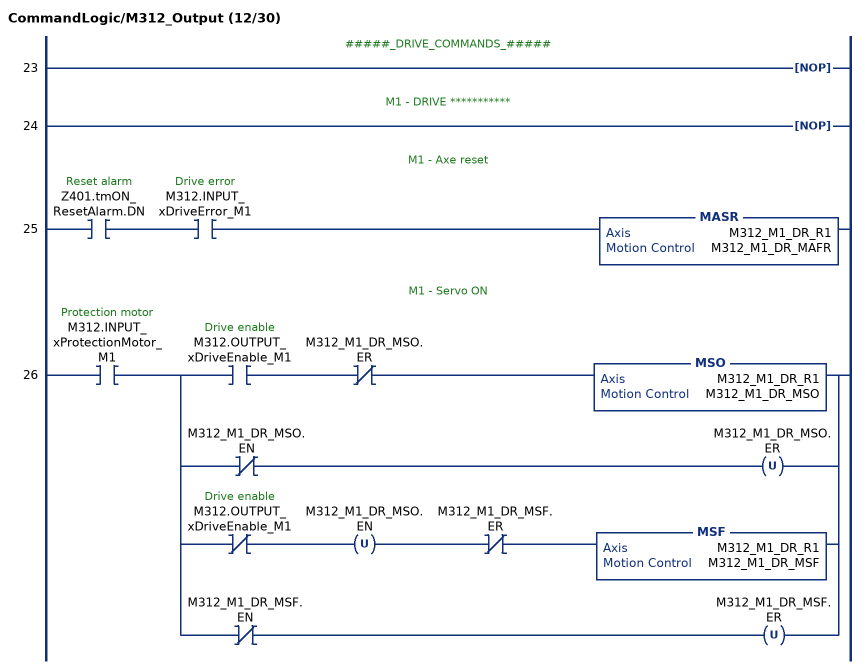
   // #####_DRIVE_COMMANDS_#####
   23: NOP();
   // M1 - DRIVE ***********
   24: NOP();
   // M1 - Axe reset
   25: XIC(Z401.tmON_ResetAlarm.DN)XIC(M312.INPUT_xDriveError_M1)MASR(M312_M1_DR_R1,M312_M1_DR_MAFR);
   // M1 - Servo ON
   26: XIC(M312.INPUT_xProtectionMotor_M1)[XIC(M312.OUTPUT_xDriveEnable_M1) XIO(M312_M1_DR_MSO.ER) MSO(M312_M1_DR_R1,M312_M1_DR_MSO) ,XIO(M312_M1_DR_MSO.EN) OTU(M312_M1_DR_MSO.ER) ,XIO(M312.OUTPUT_xDriveEnable_M1) OTU(M312_M1_DR_MSO.EN) XIO(M312_M1_DR_MSF.ER) MSF(M312_M1_DR_R1,M312_M1_DR_MSF) ,XIO(M312_M1_DR_MSF.EN) OTU(M312_M1_DR_MSF.ER) ];
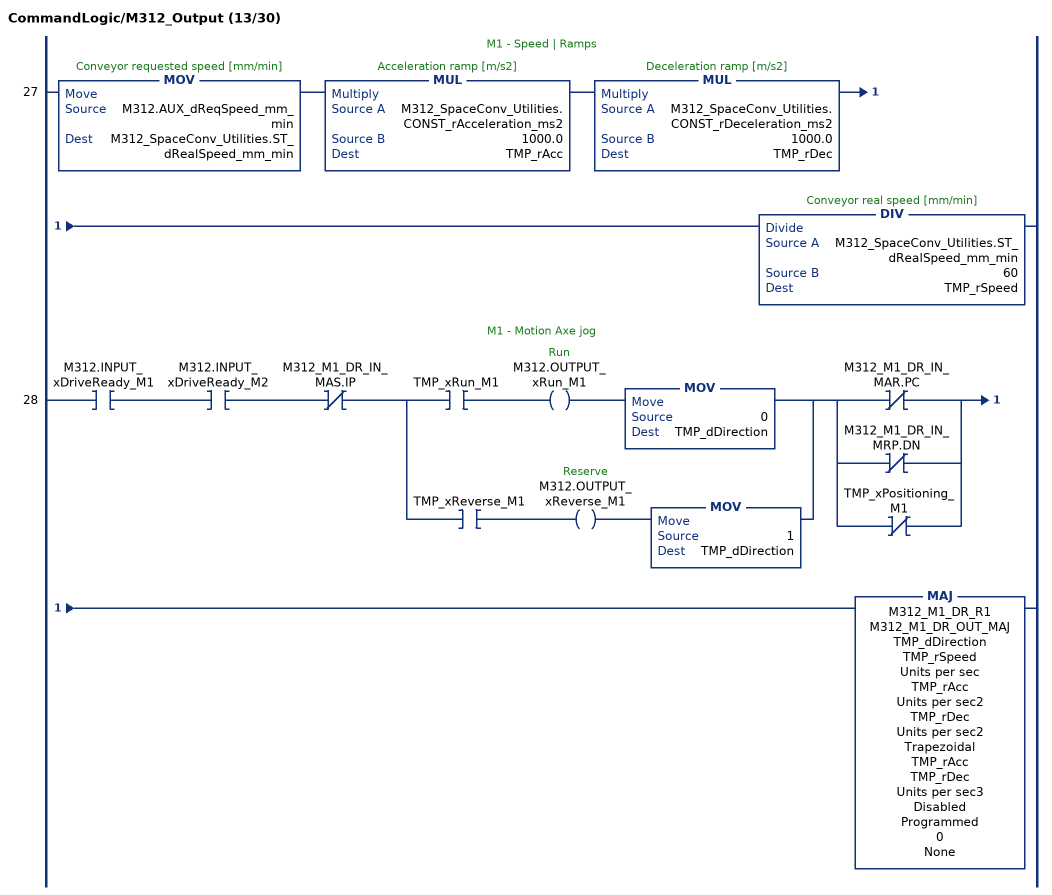
   // M1 - Speed | Ramps
   27: MOV(M312.AUX_dReqSpeed_mm_min,M312_SpaceConv_Utilities.ST_dRealSpeed_mm_min)MUL(M312_SpaceConv_Utilities.CONST_rAcceleration_ms2,1000.0,TMP_rAcc)MUL(M312_SpaceConv_Utilities.CONST_rDeceleration_ms2,1000.0,TMP_rDec)DIV(M312_SpaceConv_Utilities.ST_dRealSpeed_mm_min,60,TMP_rSpeed);
   // M1 - Motion Axe jog
   28: XIC(M312.INPUT_xDriveReady_M1)XIC(M312.INPUT_xDriveReady_M2)XIO(M312_M1_DR_IN_MAS.IP)[XIC(TMP_xRun_M1) OTE(M312.OUTPUT_xRun_M1) MOV(0,TMP_dDirection) ,XIC(TMP_xReverse_M1) OTE(M312.OUTPUT_xReverse_M1) MOV(1,TMP_dDirection) ][XIO(M312_M1_DR_IN_MAR.PC) ,XIO(M312_M1_DR_IN_MRP.DN) ,XIO(TMP_xPositioning_M1) ]MAJ(M312_M1_DR_R1,M312_M1_DR_OUT_MAJ,TMP_dDirection,TMP_rSpeed,Units per sec,TMP_rAcc,Units per sec2,TMP_rDec,Units per sec2,Trapezoidal,TMP_rAcc,TMP_rDec,Units per sec3,Disabled,Programmed,0,None);
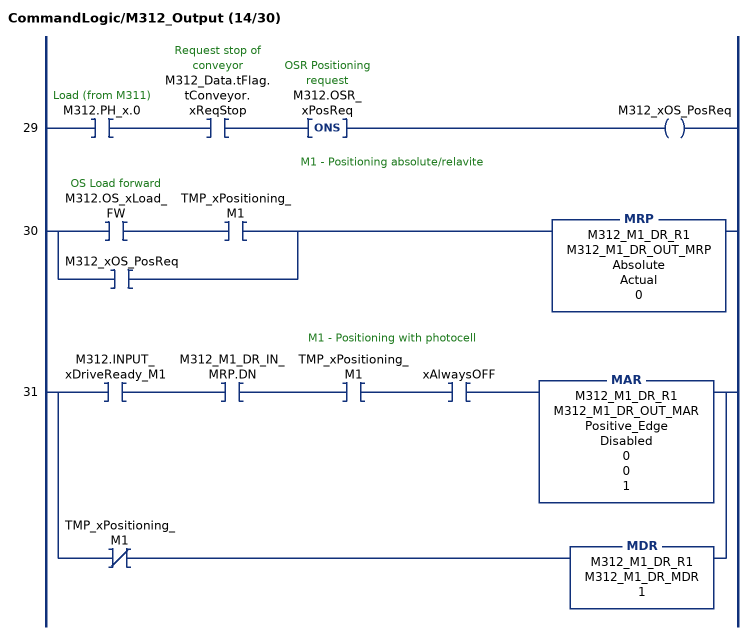
   29: XIC(M312.PH_x.0)XIC(M312_Data.tFlag.tConveyor.xReqStop)ONS(M312.OSR_xPosReq)OTE(M312_xOS_PosReq);
   // M1 - Positioning absolute/relavite
   30: [XIC(M312.OS_xLoad_FW) XIC(TMP_xPositioning_M1) ,XIC(M312_xOS_PosReq) ]MRP(M312_M1_DR_R1,M312_M1_DR_OUT_MRP,Absolute,Actual,0);
   // M1 - Positioning with photocell
   31: [XIC(M312.INPUT_xDriveReady_M1) XIC(M312_M1_DR_IN_MRP.DN) XIC(TMP_xPositioning_M1) XIC(xAlwaysOFF) MAR(M312_M1_DR_R1,M312_M1_DR_OUT_MAR,Positive_Edge,Disabled,0,0,1) ,XIO(TMP_xPositioning_M1) MDR(M312_M1_DR_R1,M312_M1_DR_MDR,1) ];
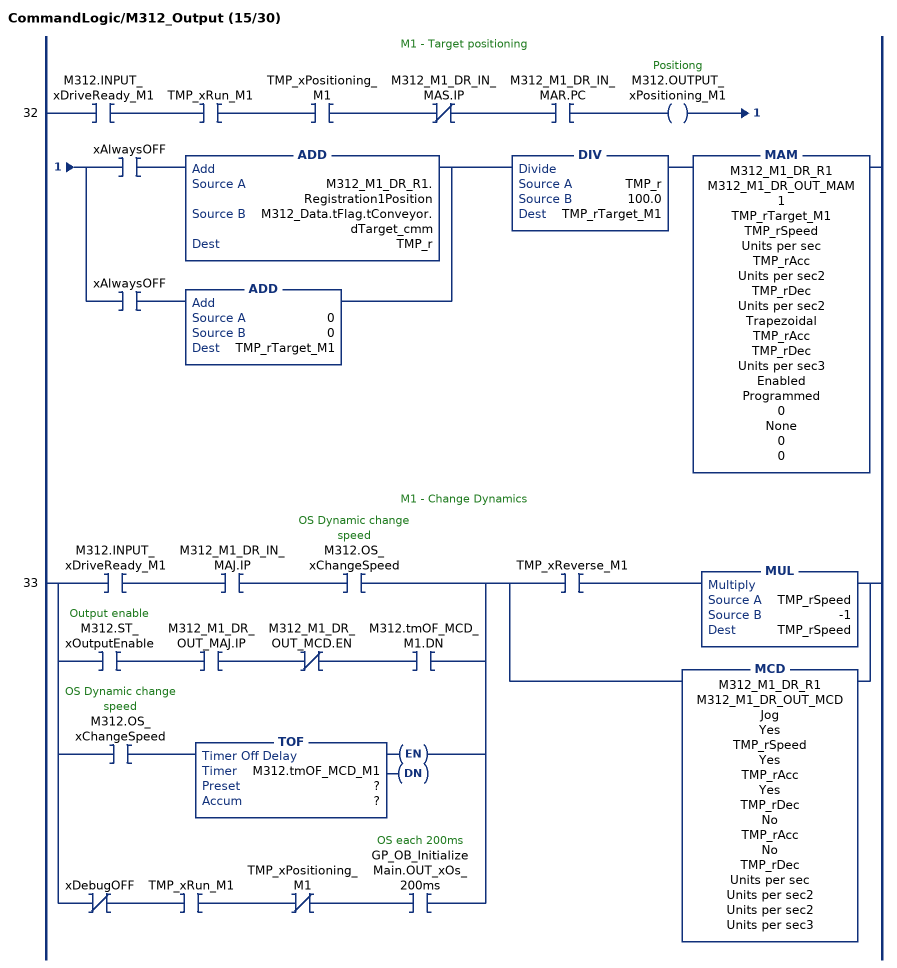
   // M1 - Target positioning
   32: XIC(M312.INPUT_xDriveReady_M1)XIC(TMP_xRun_M1)XIC(TMP_xPositioning_M1)XIO(M312_M1_DR_IN_MAS.IP)XIC(M312_M1_DR_IN_MAR.PC)OTE(M312.OUTPUT_xPositioning_M1)[XIC(xAlwaysOFF) ADD(M312_M1_DR_R1.Registration1Position,M312_Data.tFlag.tConveyor.dTarget_cmm,TMP_r) ,XIC(xAlwaysOFF) ADD(0,0,TMP_rTarget_M1) ]DIV(TMP_r,100.0,TMP_rTarget_M1)MAM(M312_M1_DR_R1,M312_M1_DR_OUT_MAM,1,TMP_rTarget_M1,TMP_rSpeed,Units per sec,TMP_rAcc,Units per sec2,TMP_rDec,Units per sec2,Trapezoidal,TMP_rAcc,TMP_rDec,Units per sec3,Enabled,Programmed,0,None,0,0);
   // M1 - Change Dynamics
   33: [XIC(M312.INPUT_xDriveReady_M1) XIC(M312_M1_DR_IN_MAJ.IP) XIC(M312.OS_xChangeSpeed) ,XIC(M312.ST_xOutputEnable) XIC(M312_M1_DR_OUT_MAJ.IP) XIO(M312_M1_DR_OUT_MCD.EN) XIC(M312.tmOF_MCD_M1.DN) ,XIC(M312.OS_xChangeSpeed) TOF(M312.tmOF_MCD_M1,?,?) ,XIO(xDebugOFF) XIC(TMP_xRun_M1) XIO(TMP_xPositioning_M1) XIC(GP_OB_InitializeMain.OUT_xOs_200ms) ][XIC(TMP_xReverse_M1) MUL(TMP_rSpeed,-1,TMP_rSpeed) ,MCD(M312_M1_DR_R1,M312_M1_DR_OUT_MCD,Jog,Yes,TMP_rSpeed,Yes,TMP_rAcc,Yes,TMP_rDec,No,TMP_rAcc,No,TMP_rDec,Units per sec,Units per sec2,Units per sec2,Units per sec3) ];
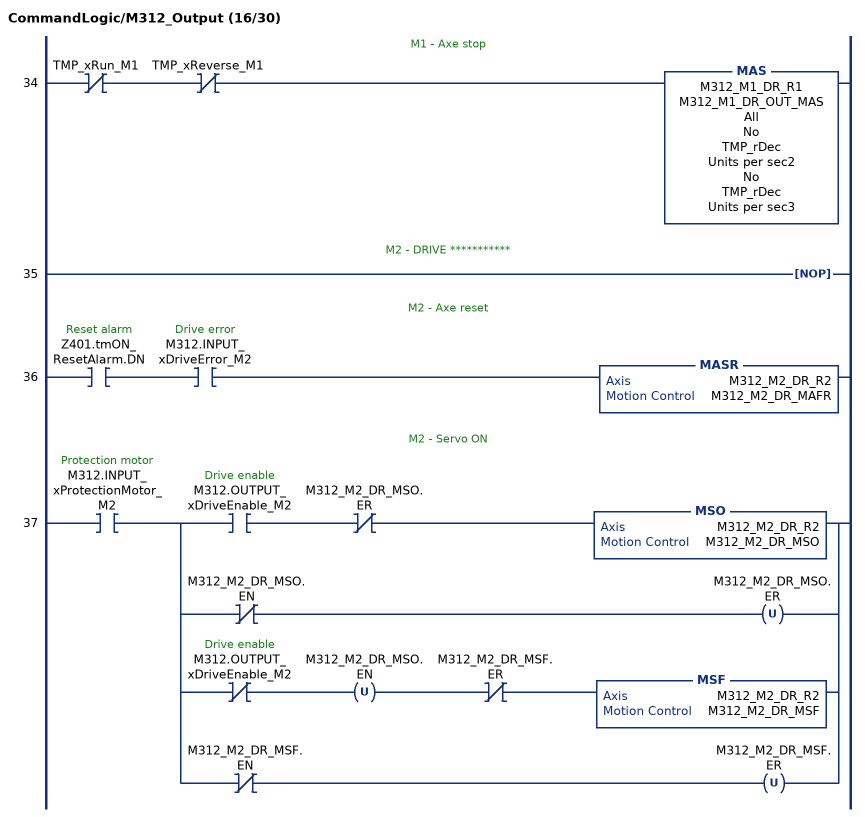
   // M1 - Axe stop
   34: XIO(TMP_xRun_M1)XIO(TMP_xReverse_M1)MAS(M312_M1_DR_R1,M312_M1_DR_OUT_MAS,All,No,TMP_rDec,Units per sec2,No,TMP_rDec,Units per sec3);
   // M2 - DRIVE ***********
   35: NOP();
   // M2 - Axe reset
   36: XIC(Z401.tmON_ResetAlarm.DN)XIC(M312.INPUT_xDriveError_M2)MASR(M312_M2_DR_R2,M312_M2_DR_MAFR);
   // M2 - Servo ON
   37: XIC(M312.INPUT_xProtectionMotor_M2)[XIC(M312.OUTPUT_xDriveEnable_M2) XIO(M312_M2_DR_MSO.ER) MSO(M312_M2_DR_R2,M312_M2_DR_MSO) ,XIO(M312_M2_DR_MSO.EN) OTU(M312_M2_DR_MSO.ER) ,XIO(M312.OUTPUT_xDriveEnable_M2) OTU(M312_M2_DR_MSO.EN) XIO(M312_M2_DR_MSF.ER) MSF(M312_M2_DR_R2,M312_M2_DR_MSF) ,XIO(M312_M2_DR_MSF.EN) OTU(M312_M2_DR_MSF.ER) ];
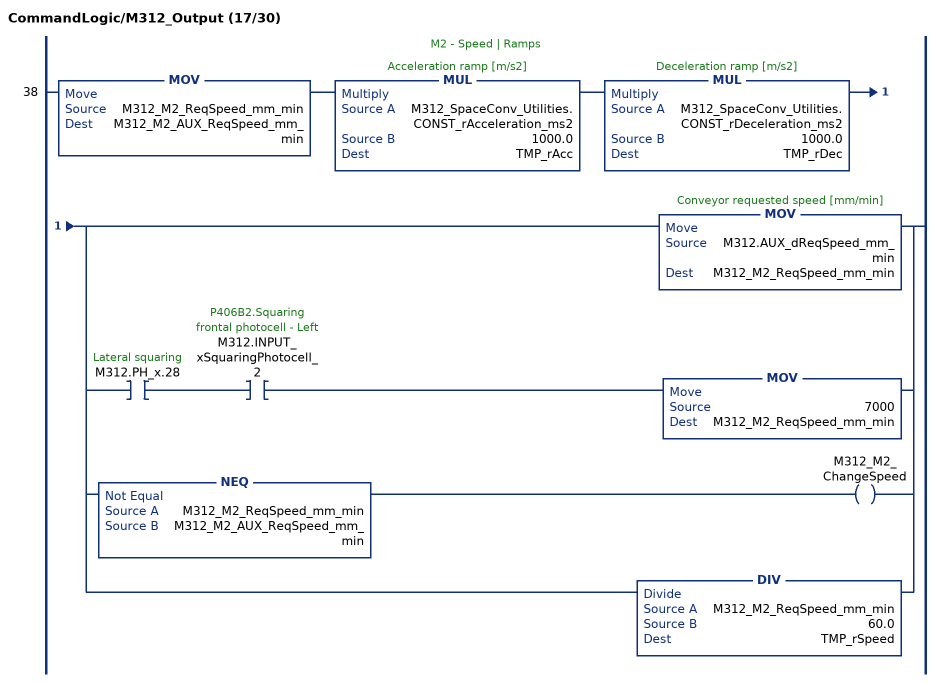
   // M2 - Speed | Ramps
   38: MOV(M312_M2_ReqSpeed_mm_min,M312_M2_AUX_ReqSpeed_mm_min)MUL(M312_SpaceConv_Utilities.CONST_rAcceleration_ms2,1000.0,TMP_rAcc)MUL(M312_SpaceConv_Utilities.CONST_rDeceleration_ms2,1000.0,TMP_rDec)[MOV(M312.AUX_dReqSpeed_mm_min,M312_M2_ReqSpeed_mm_min) ,XIC(M312.PH_x.28) XIC(M312.INPUT_xSquaringPhotocell_2) MOV(7000,M312_M2_ReqSpeed_mm_min) ,NEQ(M312_M2_ReqSpeed_mm_min,M312_M2_AUX_ReqSpeed_mm_min) OTE(M312_M2_ChangeSpeed) ,DIV(M312_M2_ReqSpeed_mm_min,60.0,TMP_rSpeed) ];
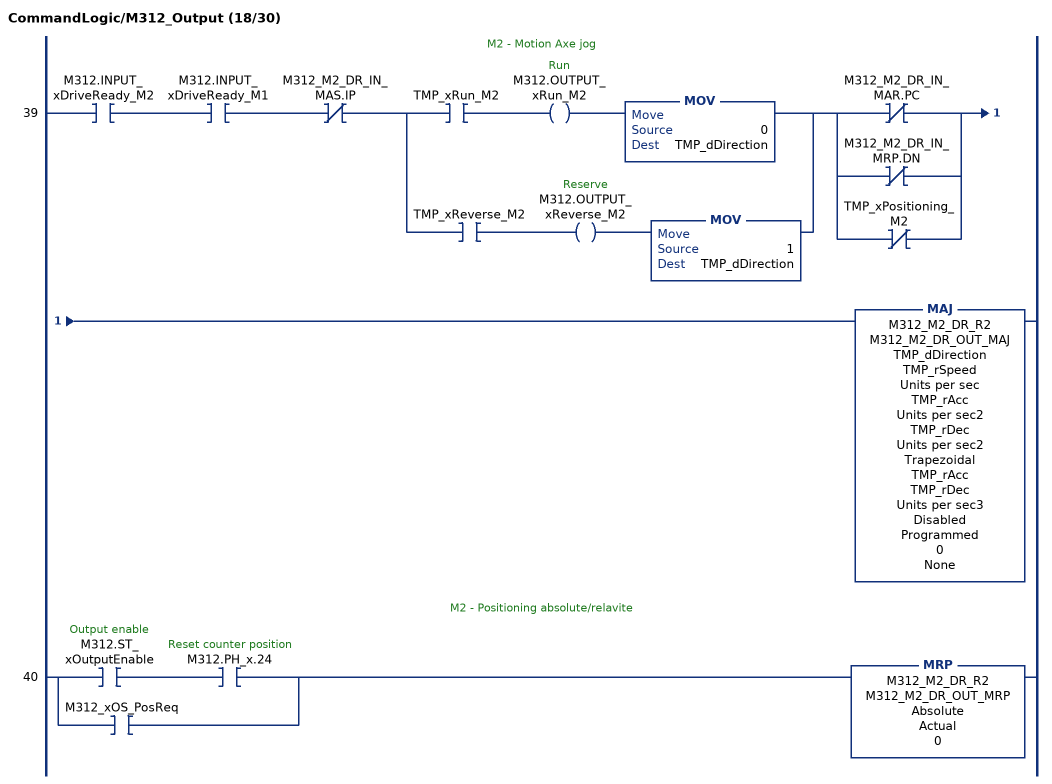
   // M2 - Motion Axe jog
   39: XIC(M312.INPUT_xDriveReady_M2)XIC(M312.INPUT_xDriveReady_M1)XIO(M312_M2_DR_IN_MAS.IP)[XIC(TMP_xRun_M2) OTE(M312.OUTPUT_xRun_M2) MOV(0,TMP_dDirection) ,XIC(TMP_xReverse_M2) OTE(M312.OUTPUT_xReverse_M2) MOV(1,TMP_dDirection) ][XIO(M312_M2_DR_IN_MAR.PC) ,XIO(M312_M2_DR_IN_MRP.DN) ,XIO(TMP_xPositioning_M2) ]MAJ(M312_M2_DR_R2,M312_M2_DR_OUT_MAJ,TMP_dDirection,TMP_rSpeed,Units per sec,TMP_rAcc,Units per sec2,TMP_rDec,Units per sec2,Trapezoidal,TMP_rAcc,TMP_rDec,Units per sec3,Disabled,Programmed,0,None);
   // M2 - Positioning absolute/relavite
   40: [XIC(M312.ST_xOutputEnable) XIC(M312.PH_x.24) ,XIC(M312_xOS_PosReq) ]MRP(M312_M2_DR_R2,M312_M2_DR_OUT_MRP,Absolute,Actual,0);
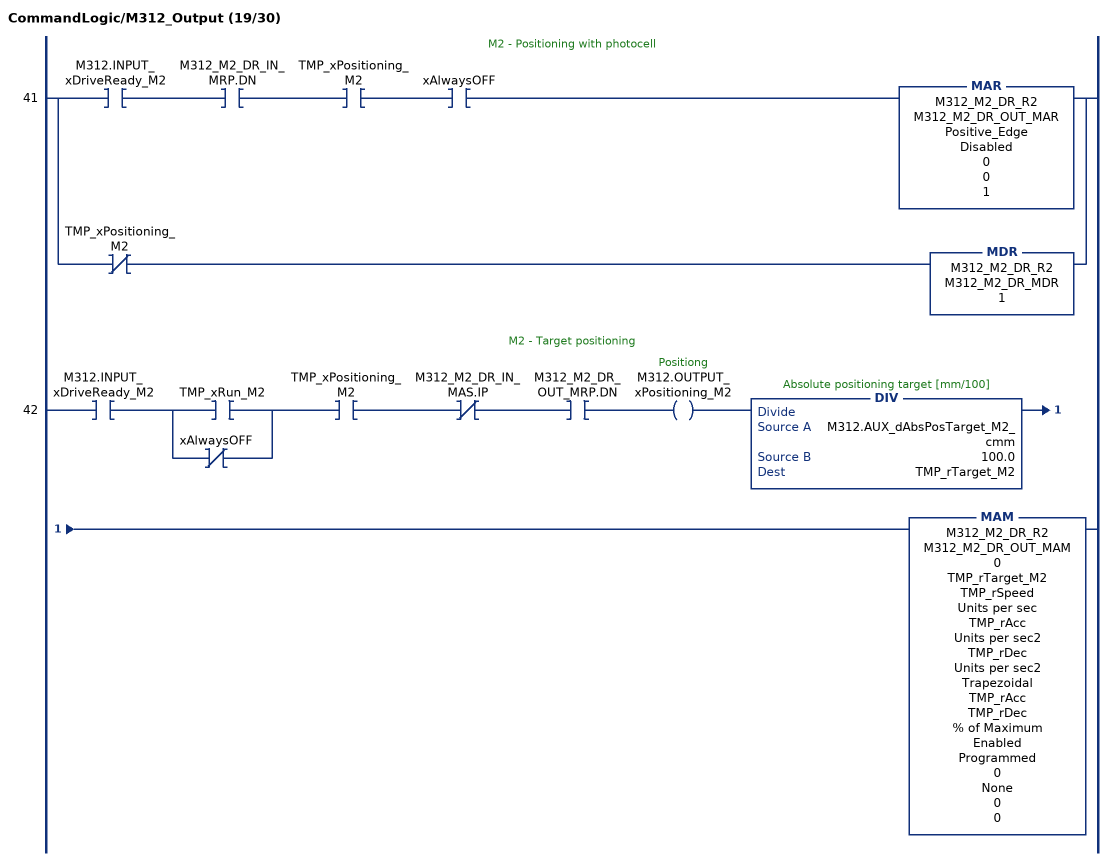
   // M2 - Positioning with photocell
   41: [XIC(M312.INPUT_xDriveReady_M2) XIC(M312_M2_DR_IN_MRP.DN) XIC(TMP_xPositioning_M2) XIC(xAlwaysOFF) MAR(M312_M2_DR_R2,M312_M2_DR_OUT_MAR,Positive_Edge,Disabled,0,0,1) ,XIO(TMP_xPositioning_M2) MDR(M312_M2_DR_R2,M312_M2_DR_MDR,1) ];
   // M2 - Target positioning
   42: XIC(M312.INPUT_xDriveReady_M2)[XIC(TMP_xRun_M2) ,XIO(xAlwaysOFF) ]XIC(TMP_xPositioning_M2)XIO(M312_M2_DR_IN_MAS.IP)XIC(M312_M2_DR_OUT_MRP.DN)OTE(M312.OUTPUT_xPositioning_M2)DIV(M312.AUX_dAbsPosTarget_M2_cmm,100.0,TMP_rTarget_M2)MAM(M312_M2_DR_R2,M312_M2_DR_OUT_MAM,0,TMP_rTarget_M2,TMP_rSpeed,Units per sec,TMP_rAcc,Units per sec2,TMP_rDec,Units per sec2,Trapezoidal,TMP_rAcc,TMP_rDec,% of Maximum,Enabled,Programmed,0,None,0,0);
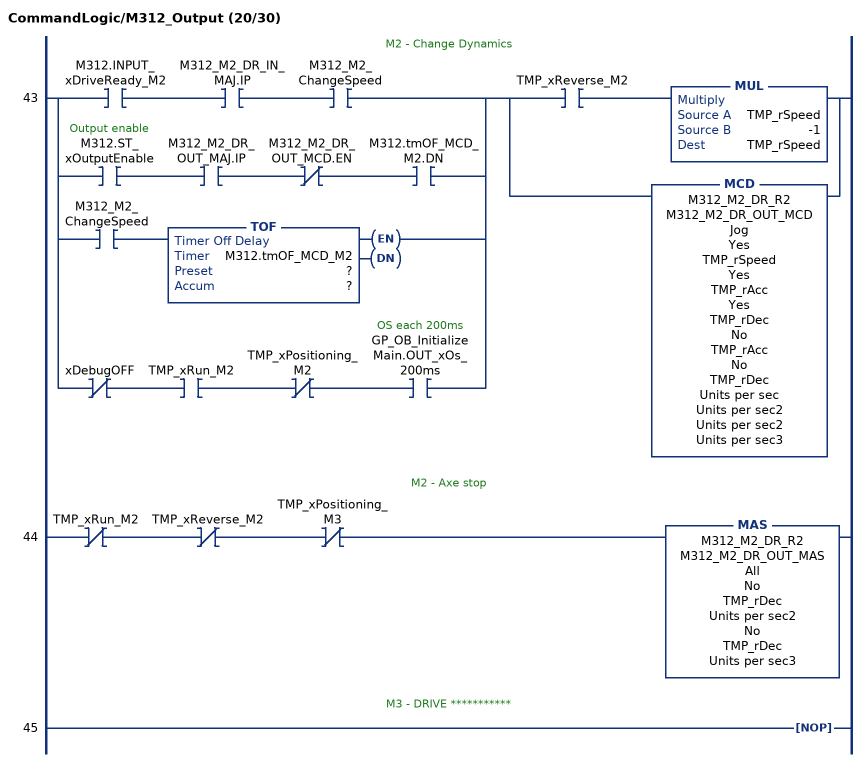
   // M2 - Change Dynamics
   43: [XIC(M312.INPUT_xDriveReady_M2) XIC(M312_M2_DR_IN_MAJ.IP) XIC(M312_M2_ChangeSpeed) ,XIC(M312.ST_xOutputEnable) XIC(M312_M2_DR_OUT_MAJ.IP) XIO(M312_M2_DR_OUT_MCD.EN) XIC(M312.tmOF_MCD_M2.DN) ,XIC(M312_M2_ChangeSpeed) TOF(M312.tmOF_MCD_M2,?,?) ,XIO(xDebugOFF) XIC(TMP_xRun_M2) XIO(TMP_xPositioning_M2) XIC(GP_OB_InitializeMain.OUT_xOs_200ms) ][XIC(TMP_xReverse_M2) MUL(TMP_rSpeed,-1,TMP_rSpeed) ,MCD(M312_M2_DR_R2,M312_M2_DR_OUT_MCD,Jog,Yes,TMP_rSpeed,Yes,TMP_rAcc,Yes,TMP_rDec,No,TMP_rAcc,No,TMP_rDec,Units per sec,Units per sec2,Units per sec2,Units per sec3) ];
   // M2 - Axe stop
   44: XIO(TMP_xRun_M2)XIO(TMP_xReverse_M2)XIO(TMP_xPositioning_M3)MAS(M312_M2_DR_R2,M312_M2_DR_OUT_MAS,All,No,TMP_rDec,Units per sec2,No,TMP_rDec,Units per sec3);
   // M3 - DRIVE ***********
   45: NOP();
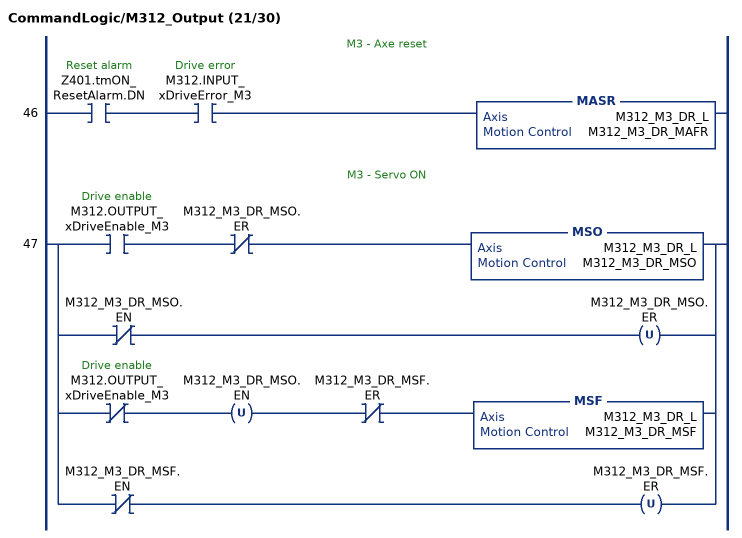
   // M3 - Axe reset
   46: XIC(Z401.tmON_ResetAlarm.DN)XIC(M312.INPUT_xDriveError_M3)MASR(M312_M3_DR_L,M312_M3_DR_MAFR);
   // M3 - Servo ON
   47: [XIC(M312.OUTPUT_xDriveEnable_M3) XIO(M312_M3_DR_MSO.ER) MSO(M312_M3_DR_L,M312_M3_DR_MSO) ,XIO(M312_M3_DR_MSO.EN) OTU(M312_M3_DR_MSO.ER) ,XIO(M312.OUTPUT_xDriveEnable_M3) OTU(M312_M3_DR_MSO.EN) XIO(M312_M3_DR_MSF.ER) MSF(M312_M3_DR_L,M312_M3_DR_MSF) ,XIO(M312_M3_DR_MSF.EN) OTU(M312_M3_DR_MSF.ER) ];
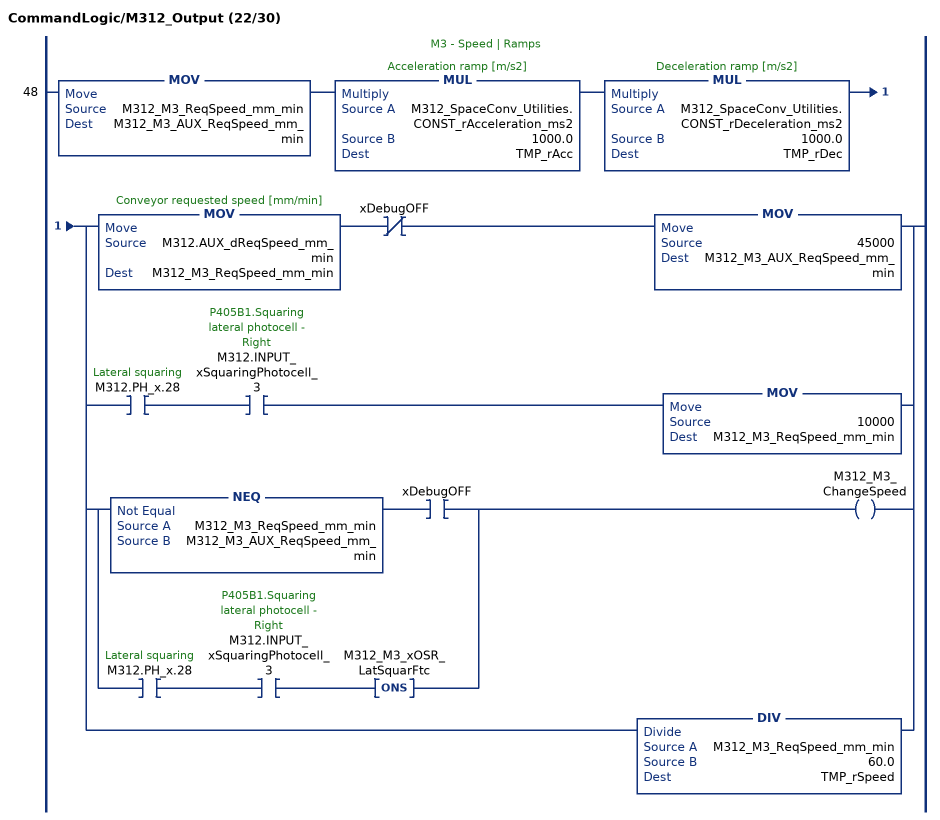
   // M3 - Speed | Ramps
   48: MOV(M312_M3_ReqSpeed_mm_min,M312_M3_AUX_ReqSpeed_mm_min)MUL(M312_SpaceConv_Utilities.CONST_rAcceleration_ms2,1000.0,TMP_rAcc)MUL(M312_SpaceConv_Utilities.CONST_rDeceleration_ms2,1000.0,TMP_rDec)[MOV(M312.AUX_dReqSpeed_mm_min,M312_M3_ReqSpeed_mm_min) XIO(xDebugOFF) MOV(45000,M312_M3_AUX_ReqSpeed_mm_min) ,XIC(M312.PH_x.28) XIC(M312.INPUT_xSquaringPhotocell_3) MOV(10000,M312_M3_ReqSpeed_mm_min) ,[NEQ(M312_M3_ReqSpeed_mm_min,M312_M3_AUX_ReqSpeed_mm_min) XIC(xDebugOFF) ,XIC(M312.PH_x.28) XIC(M312.INPUT_xSquaringPhotocell_3) ONS(M312_M3_xOSR_LatSquarFtc) ] OTE(M312_M3_ChangeSpeed) ,DIV(M312_M3_ReqSpeed_mm_min,60.0,TMP_rSpeed) ];
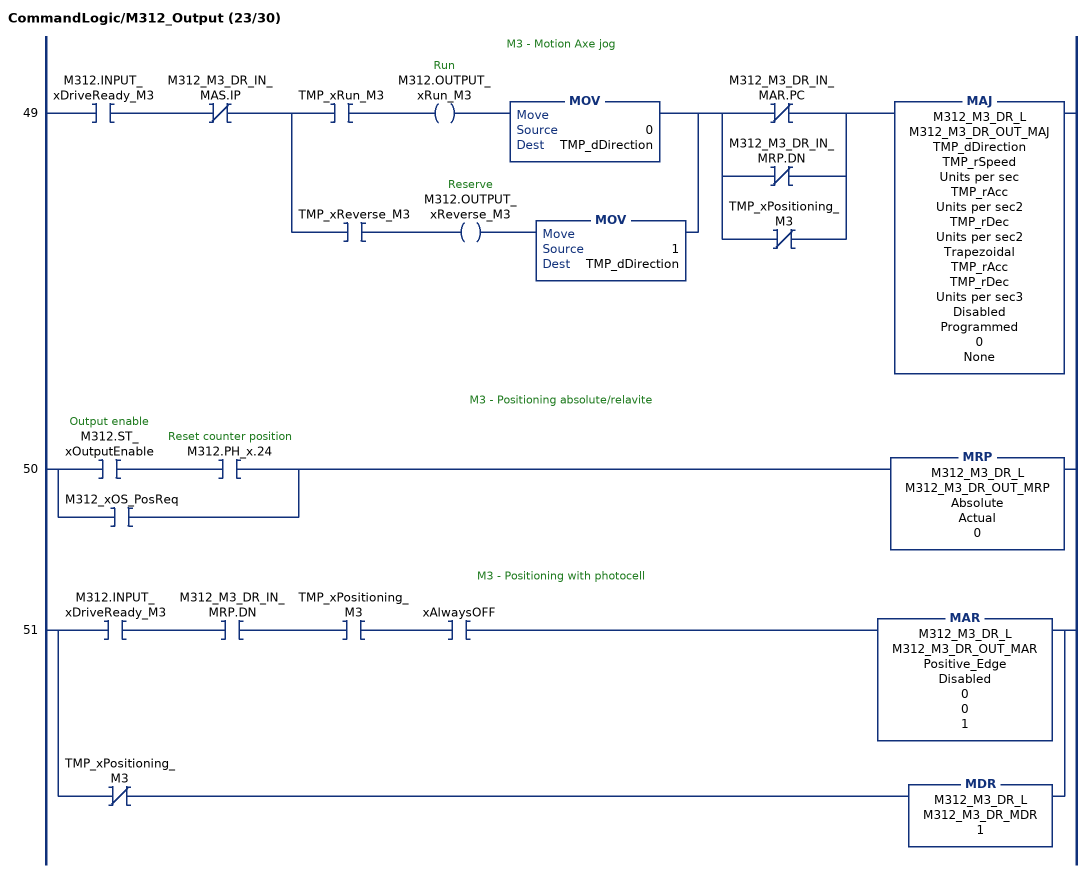
   // M3 - Motion Axe jog
   49: XIC(M312.INPUT_xDriveReady_M3)XIO(M312_M3_DR_IN_MAS.IP)[XIC(TMP_xRun_M3) OTE(M312.OUTPUT_xRun_M3) MOV(0,TMP_dDirection) ,XIC(TMP_xReverse_M3) OTE(M312.OUTPUT_xReverse_M3) MOV(1,TMP_dDirection) ][XIO(M312_M3_DR_IN_MAR.PC) ,XIO(M312_M3_DR_IN_MRP.DN) ,XIO(TMP_xPositioning_M3) ]MAJ(M312_M3_DR_L,M312_M3_DR_OUT_MAJ,TMP_dDirection,TMP_rSpeed,Units per sec,TMP_rAcc,Units per sec2,TMP_rDec,Units per sec2,Trapezoidal,TMP_rAcc,TMP_rDec,Units per sec3,Disabled,Programmed,0,None);
   // M3 - Positioning absolute/relavite
   50: [XIC(M312.ST_xOutputEnable) XIC(M312.PH_x.24) ,XIC(M312_xOS_PosReq) ]MRP(M312_M3_DR_L,M312_M3_DR_OUT_MRP,Absolute,Actual,0);
   // M3 - Positioning with photocell
   51: [XIC(M312.INPUT_xDriveReady_M3) XIC(M312_M3_DR_IN_MRP.DN) XIC(TMP_xPositioning_M3) XIC(xAlwaysOFF) MAR(M312_M3_DR_L,M312_M3_DR_OUT_MAR,Positive_Edge,Disabled,0,0,1) ,XIO(TMP_xPositioning_M3) MDR(M312_M3_DR_L,M312_M3_DR_MDR,1) ];
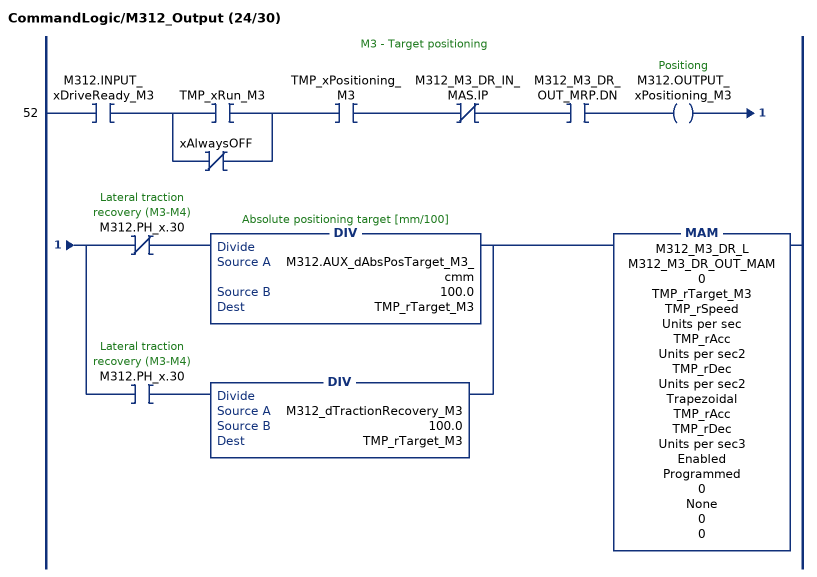
   // M3 - Target positioning
   52: XIC(M312.INPUT_xDriveReady_M3)[XIC(TMP_xRun_M3) ,XIO(xAlwaysOFF) ]XIC(TMP_xPositioning_M3)XIO(M312_M3_DR_IN_MAS.IP)XIC(M312_M3_DR_OUT_MRP.DN)OTE(M312.OUTPUT_xPositioning_M3)[XIO(M312.PH_x.30) DIV(M312.AUX_dAbsPosTarget_M3_cmm,100.0,TMP_rTarget_M3) ,XIC(M312.PH_x.30) DIV(M312_dTractionRecovery_M3,100.0,TMP_rTarget_M3) ]MAM(M312_M3_DR_L,M312_M3_DR_OUT_MAM,0,TMP_rTarget_M3,TMP_rSpeed,Units per sec,TMP_rAcc,Units per sec2,TMP_rDec,Units per sec2,Trapezoidal,TMP_rAcc,TMP_rDec,Units per sec3,Enabled,Programmed,0,None,0,0);
